// TIA Portal project "ESTHER_Gas_v4.0_4" (V13) (continued)
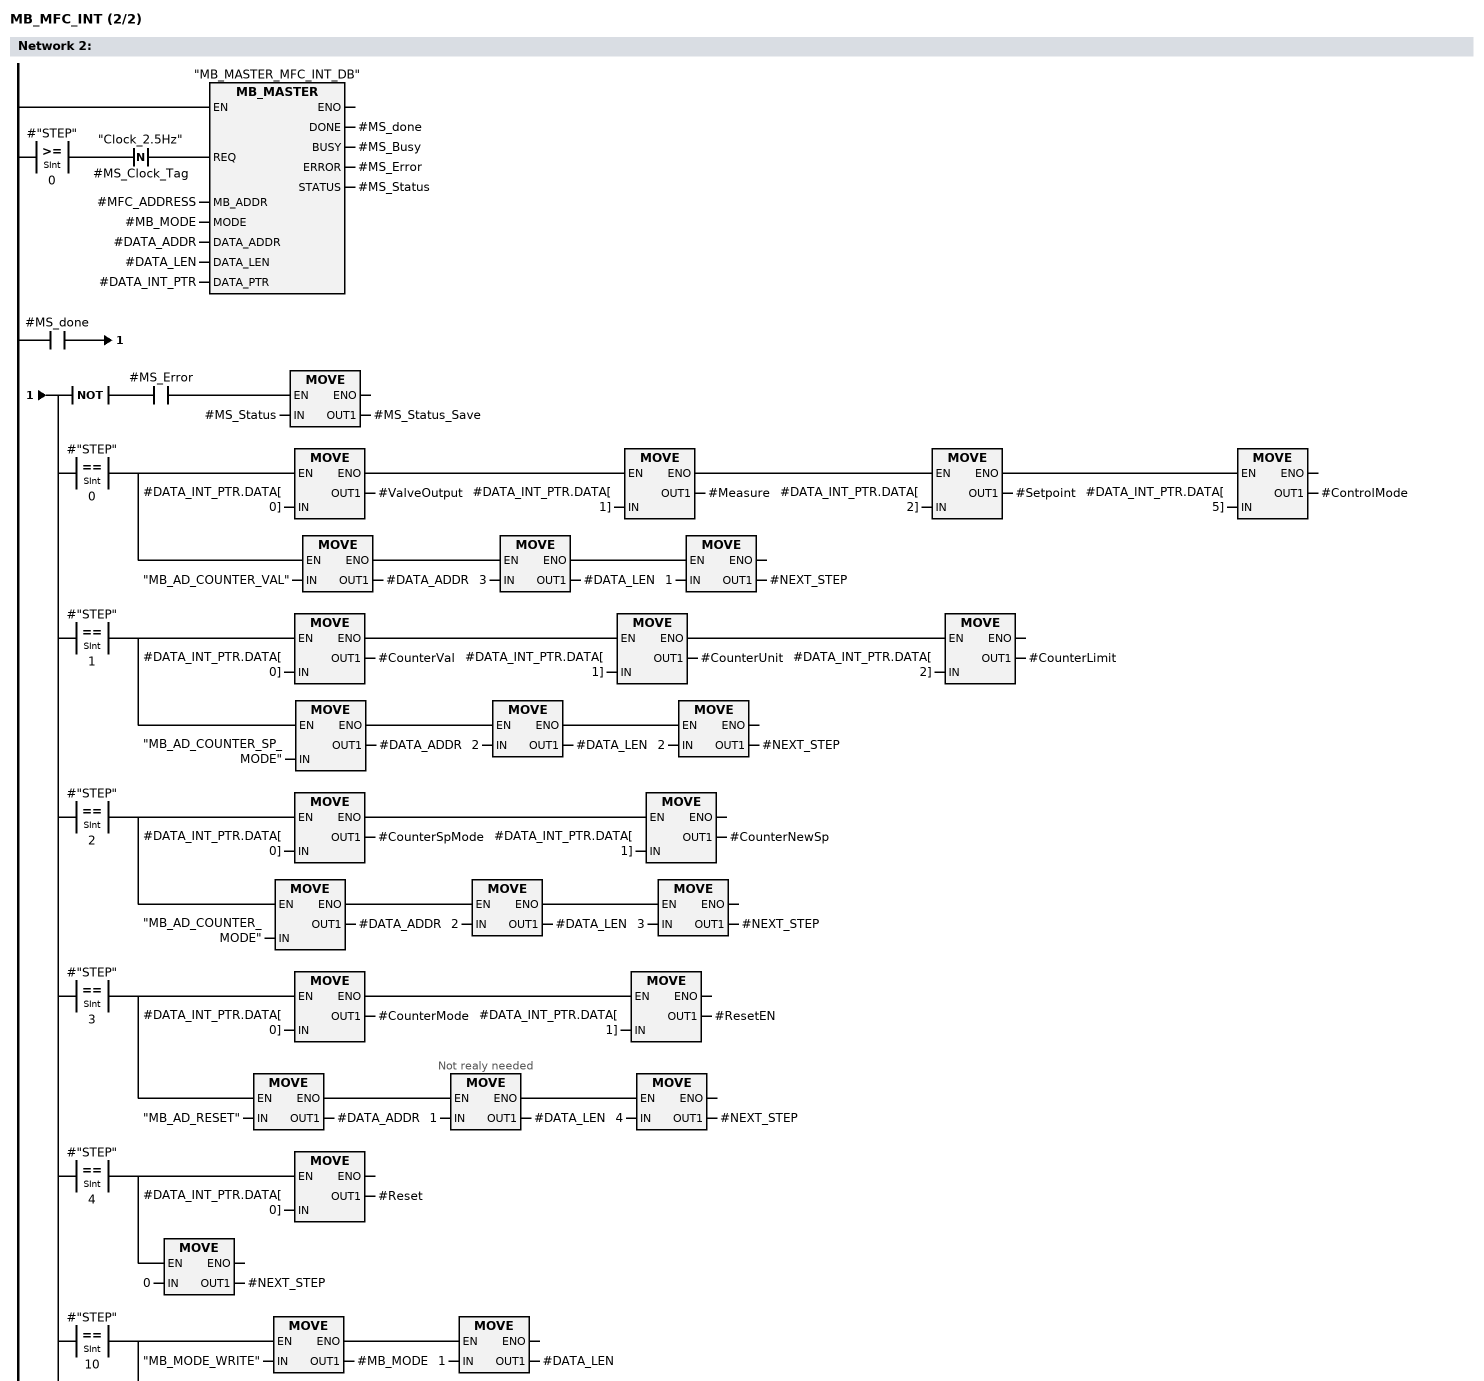
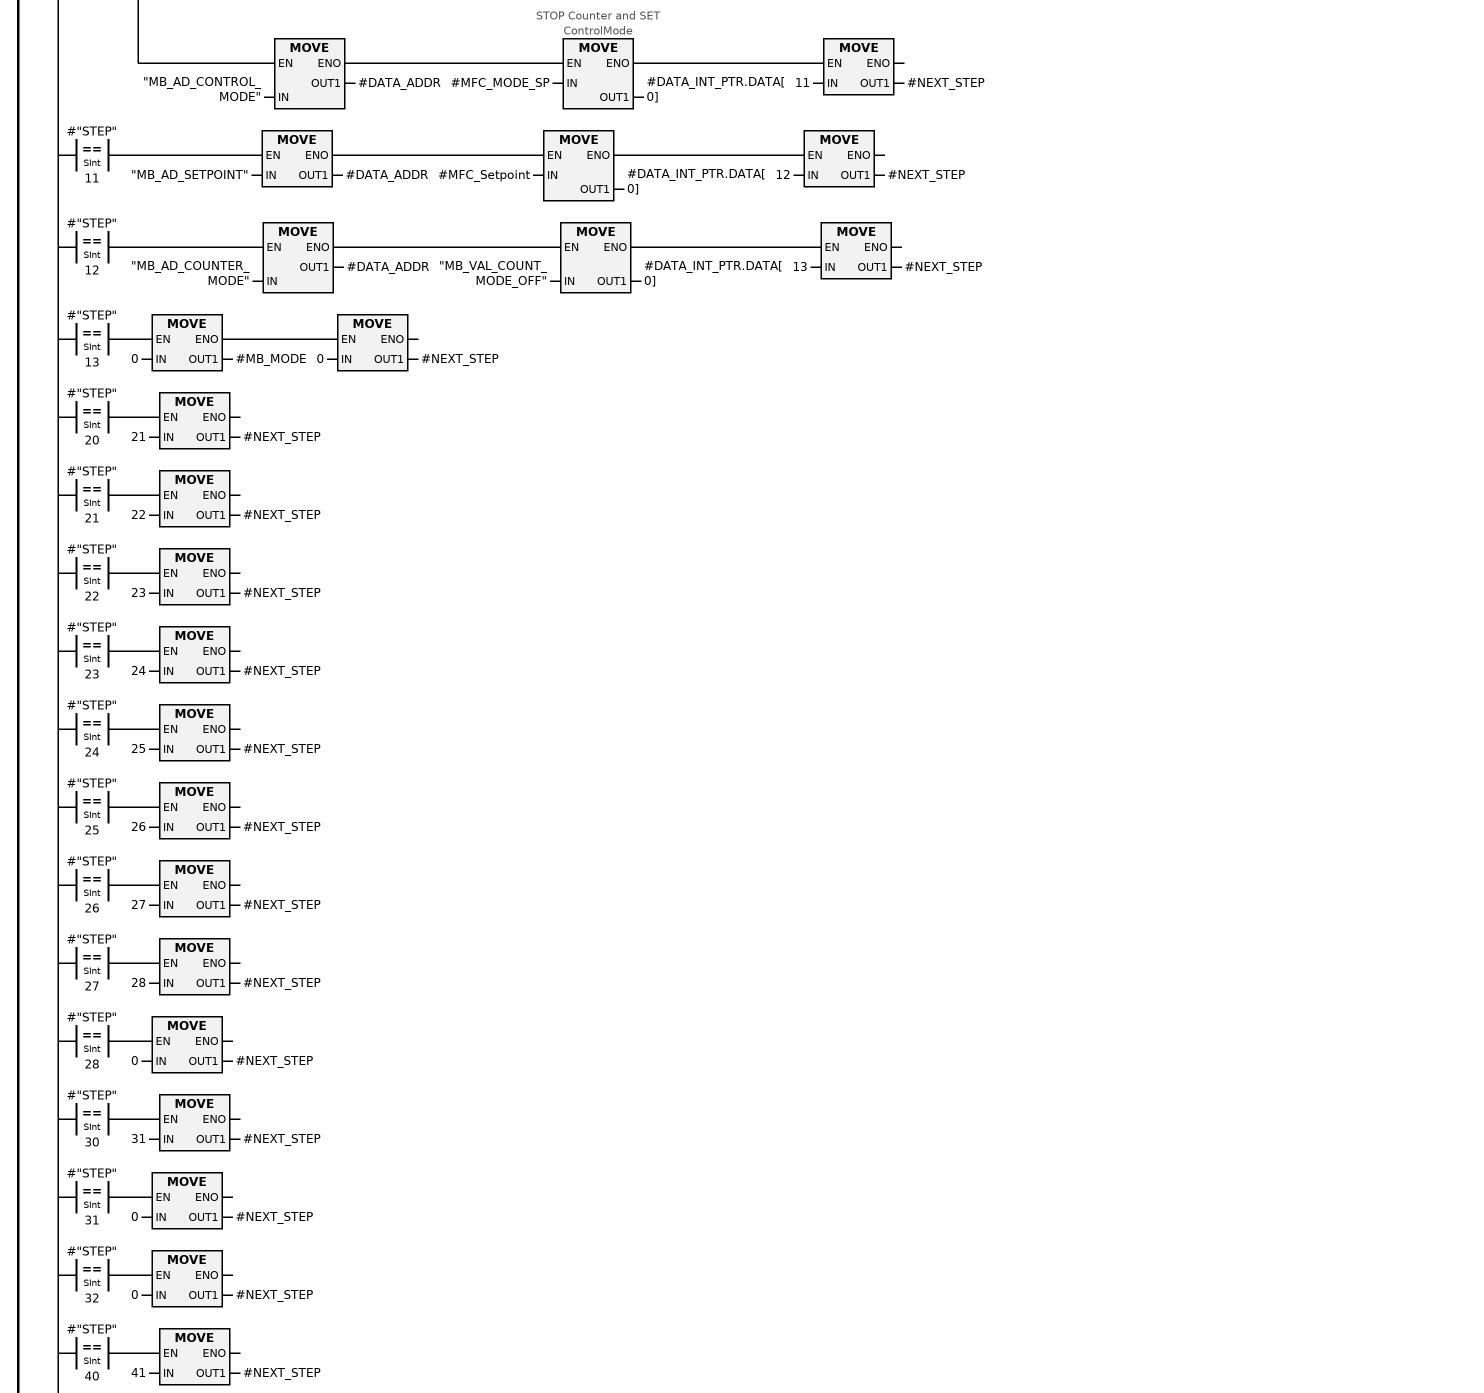
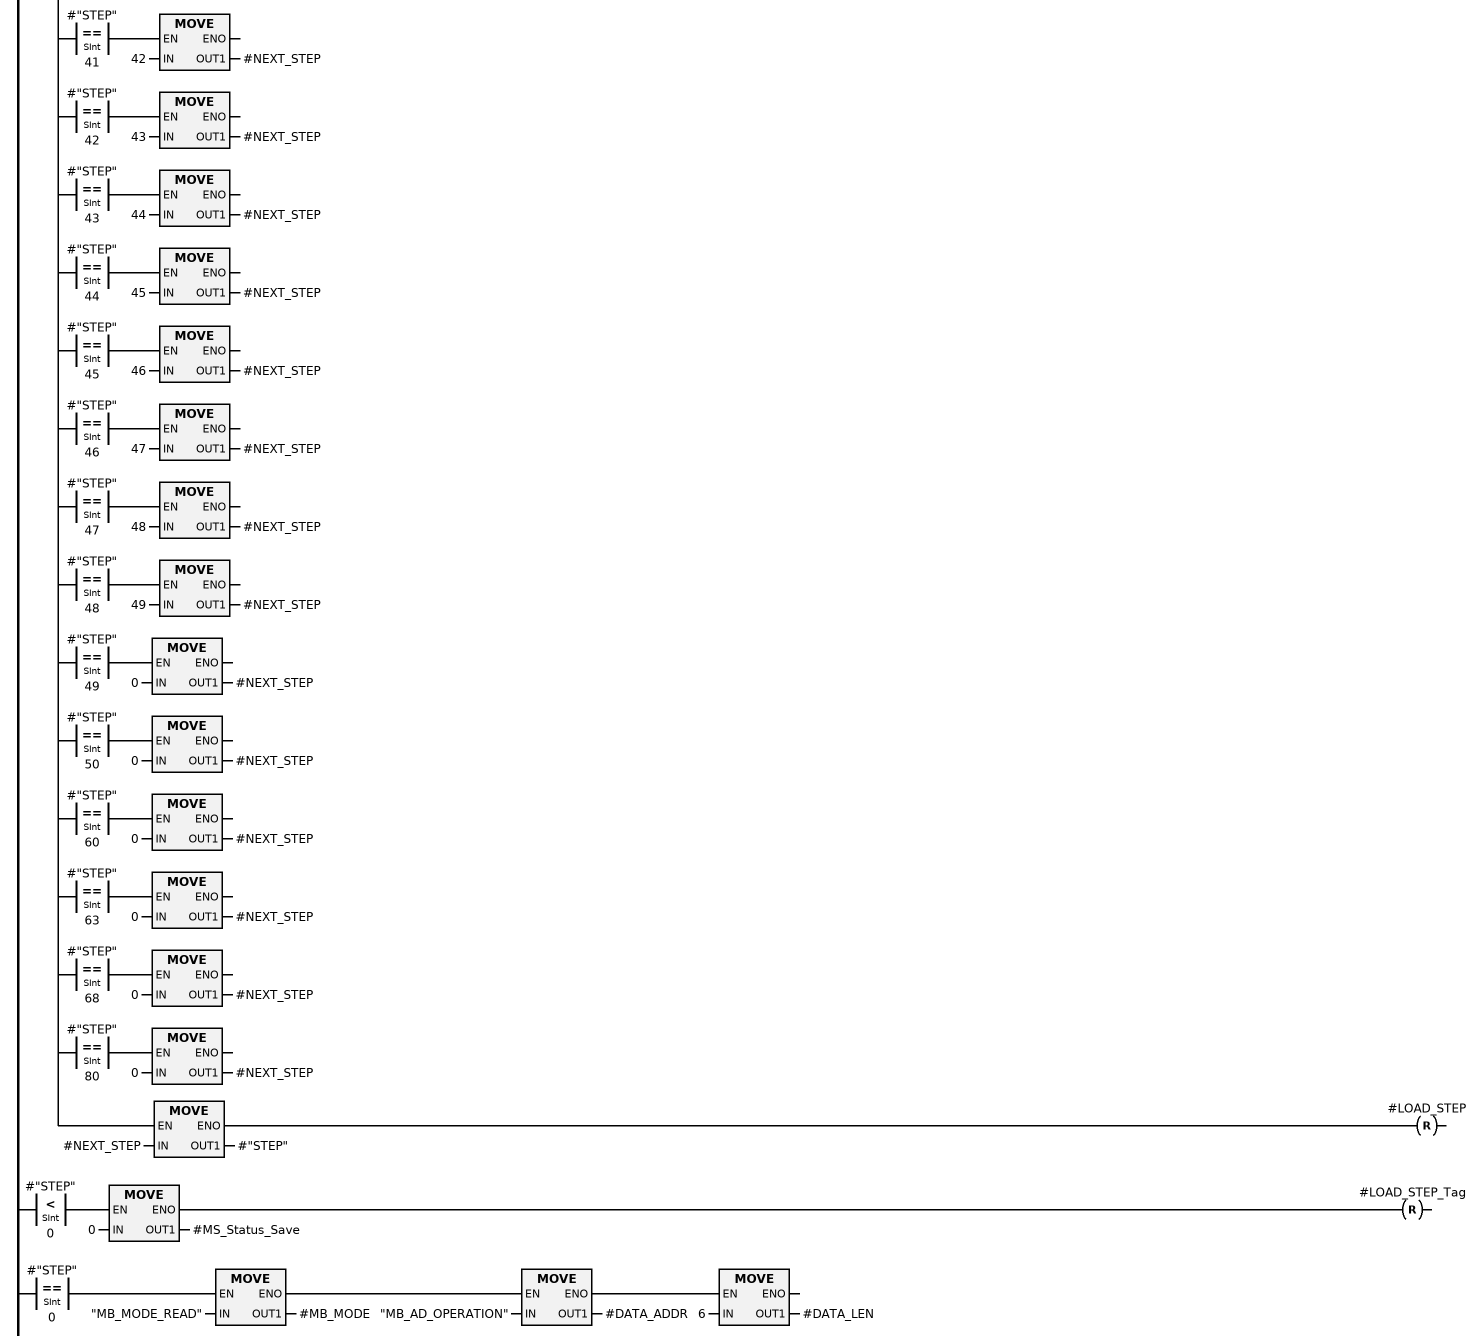
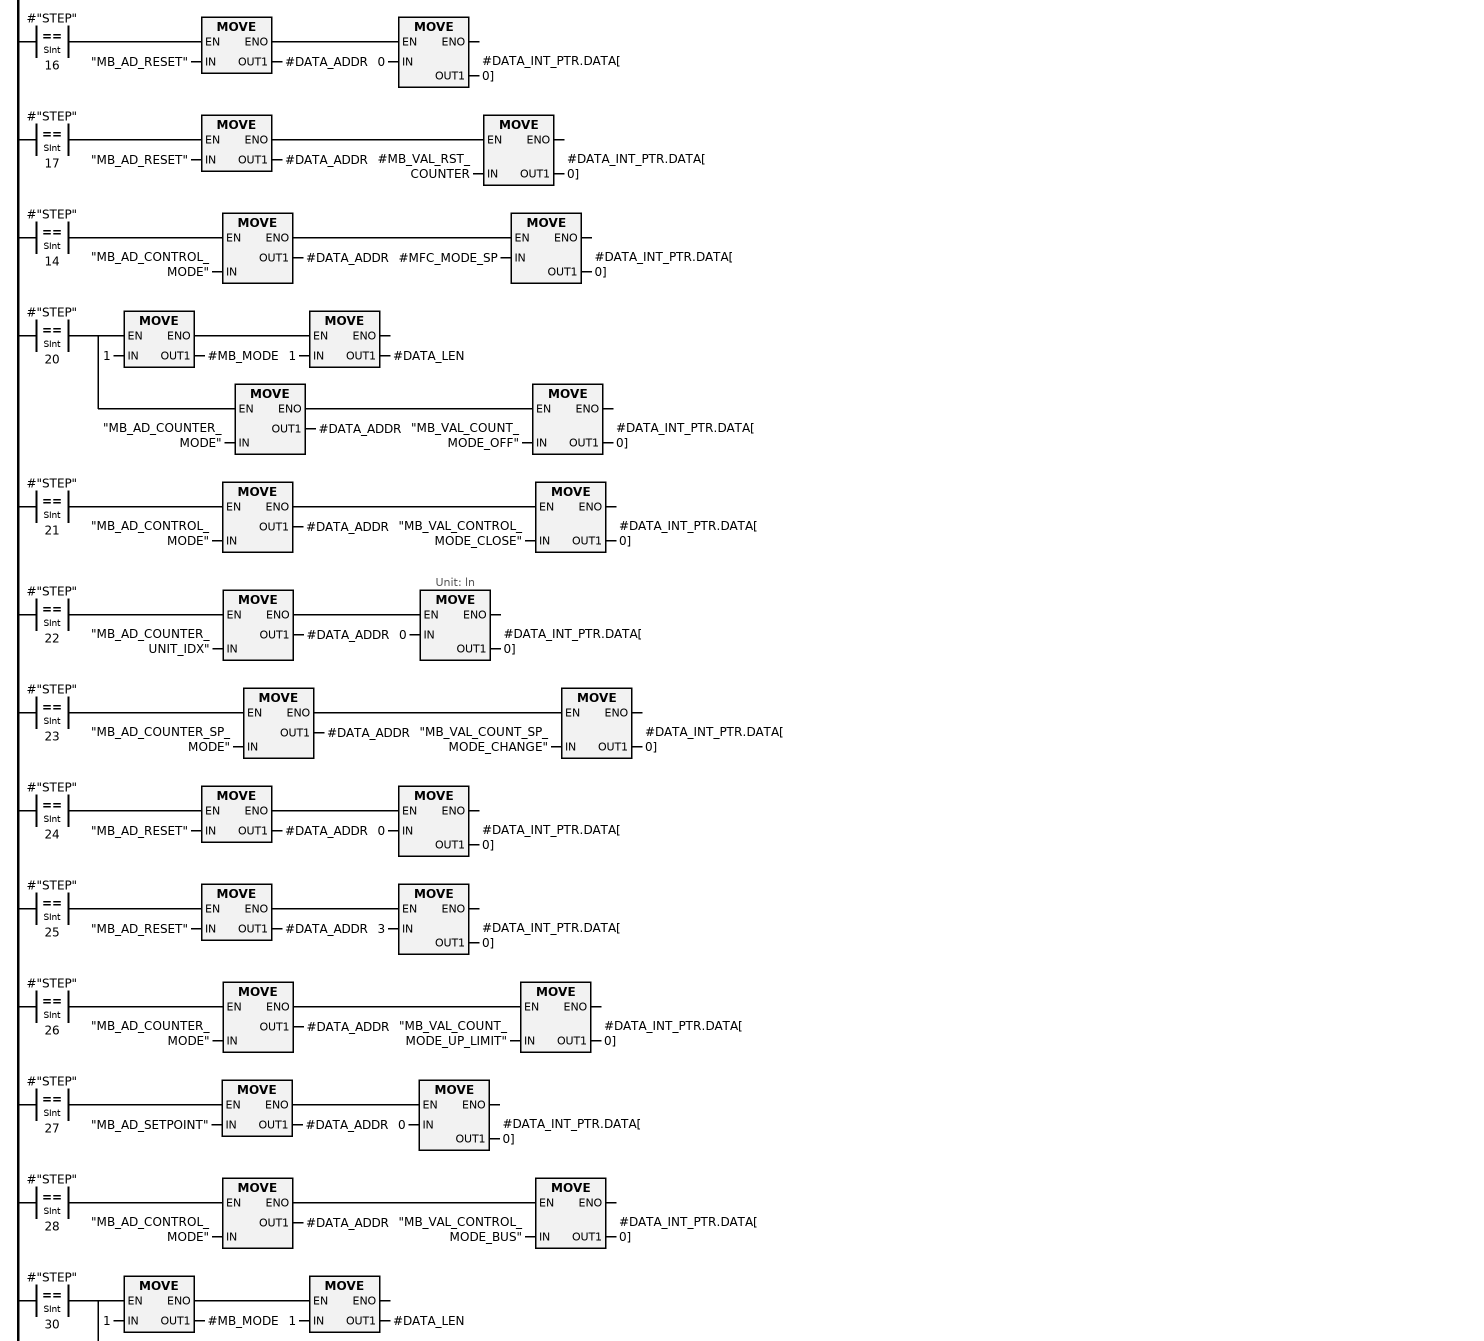
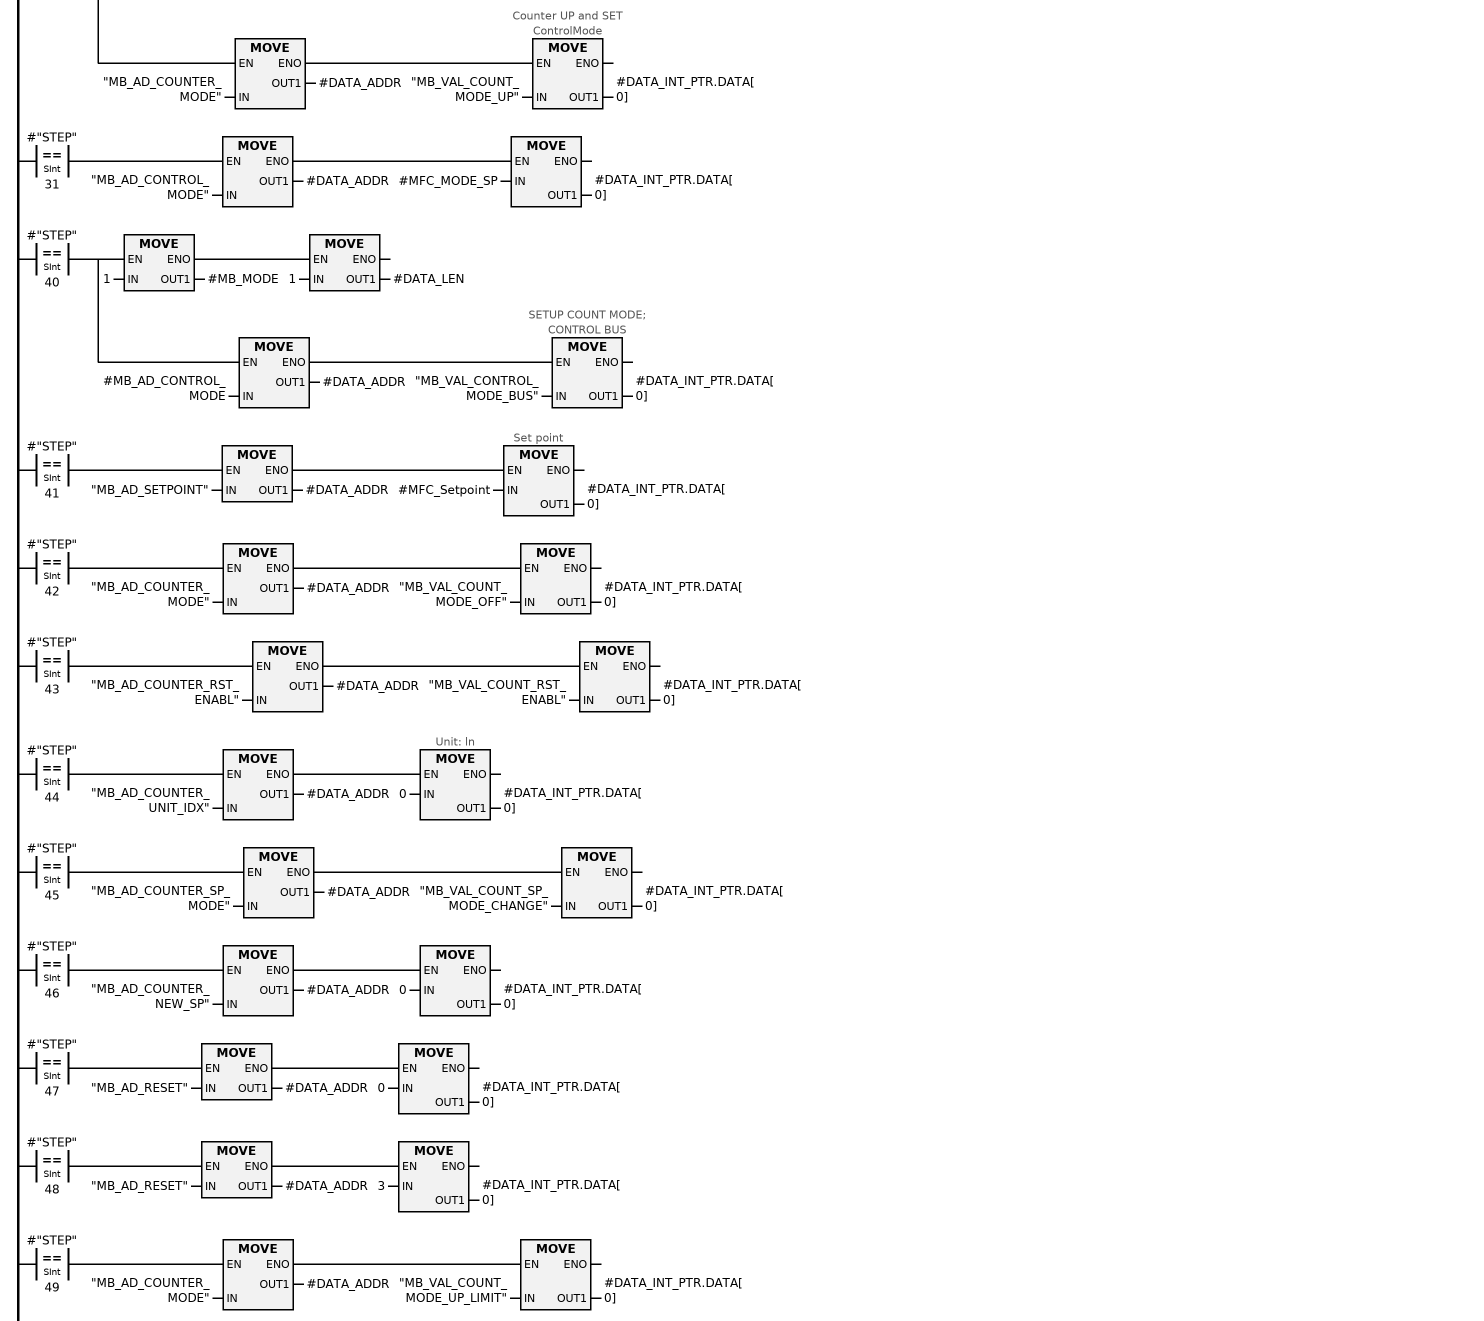
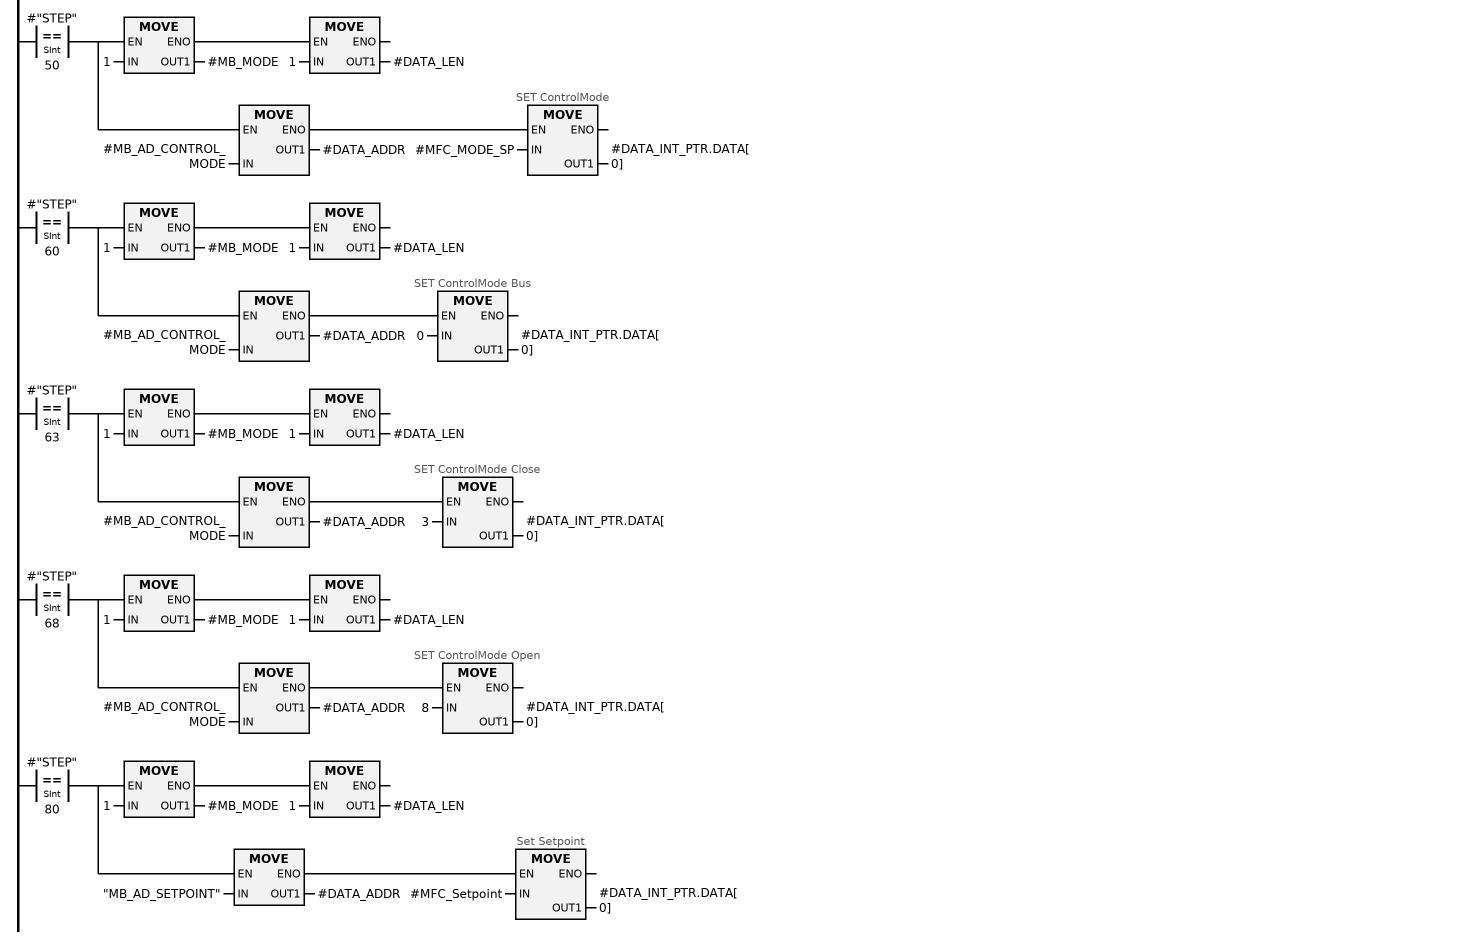
   #_w1 := (#"STEP" >= 0) AND NOT "Clock_2.5Hz" AND #MS_Clock_Tag;   // falling edge of "Clock_2.5Hz"
   #MS_Clock_Tag := "Clock_2.5Hz";
   "MB_MASTER_MFC_INT_DB"(REQ := #_w1,   // MB_MASTER
                          MB_ADDR := #MFC_ADDRESS,
                          MODE := #MB_MODE,
                          DATA_ADDR := #DATA_ADDR,
                          DATA_LEN := #DATA_LEN,
                          DATA_PTR := #DATA_INT_PTR,
                          DONE => #MS_done,
                          BUSY => #MS_Busy,
                          ERROR => #MS_Error,
                          STATUS => #MS_Status);
   IF NOT #MS_done AND #MS_Error THEN #MS_Status_Save := #MS_Status; END_IF;
   IF #MS_done AND (#"STEP" = 0) THEN
       #ValveOutput := #DATA_INT_PTR.DATA[0];
       #Measure := #DATA_INT_PTR.DATA[1];
       #Setpoint := #DATA_INT_PTR.DATA[2];
       #ControlMode := #DATA_INT_PTR.DATA[5];
       #DATA_ADDR := "MB_AD_COUNTER_VAL";
       #DATA_LEN := 3;
       #NEXT_STEP := 1;
   END_IF;
   IF #MS_done AND (#"STEP" = 1) THEN
       #CounterVal := #DATA_INT_PTR.DATA[0];
       #CounterUnit := #DATA_INT_PTR.DATA[1];
       #CounterLimit := #DATA_INT_PTR.DATA[2];
       #DATA_ADDR := "MB_AD_COUNTER_SP_MODE";
       #DATA_LEN := 2;
       #NEXT_STEP := 2;
   END_IF;
   IF #MS_done AND (#"STEP" = 2) THEN
       #CounterSpMode := #DATA_INT_PTR.DATA[0];
       #CounterNewSp := #DATA_INT_PTR.DATA[1];
       #DATA_ADDR := "MB_AD_COUNTER_MODE";
       #DATA_LEN := 2;
       #NEXT_STEP := 3;
   END_IF;
   IF #MS_done AND (#"STEP" = 3) THEN
       #CounterMode := #DATA_INT_PTR.DATA[0];
       #ResetEN := #DATA_INT_PTR.DATA[1];
       #DATA_ADDR := "MB_AD_RESET";
       #DATA_LEN := 1;   // Not realy needed
       #NEXT_STEP := 4;
   END_IF;
   IF #MS_done AND (#"STEP" = 4) THEN
       #Reset := #DATA_INT_PTR.DATA[0];
       #NEXT_STEP := 0;
   END_IF;
   IF #MS_done AND (#"STEP" = 10) THEN
       #MB_MODE := "MB_MODE_WRITE";
       #DATA_LEN := 1;
       #DATA_ADDR := "MB_AD_CONTROL_MODE";
       #DATA_INT_PTR.DATA[0] := #MFC_MODE_SP;   // STOP Counter and SET ControlMode
       #NEXT_STEP := 11;
   END_IF;
   IF #MS_done AND (#"STEP" = 11) THEN
       #DATA_ADDR := "MB_AD_SETPOINT";
       #DATA_INT_PTR.DATA[0] := #MFC_Setpoint;
       #NEXT_STEP := 12;
   END_IF;
   IF #MS_done AND (#"STEP" = 12) THEN
       #DATA_ADDR := "MB_AD_COUNTER_MODE";
       #DATA_INT_PTR.DATA[0] := "MB_VAL_COUNT_MODE_OFF";
       #NEXT_STEP := 13;
   END_IF;
   IF #MS_done AND (#"STEP" = 13) THEN
       #MB_MODE := 0;
       #NEXT_STEP := 0;
   END_IF;
   IF #MS_done AND (#"STEP" = 20) THEN #NEXT_STEP := 21; END_IF;
   IF #MS_done AND (#"STEP" = 21) THEN #NEXT_STEP := 22; END_IF;
   IF #MS_done AND (#"STEP" = 22) THEN #NEXT_STEP := 23; END_IF;
   IF #MS_done AND (#"STEP" = 23) THEN #NEXT_STEP := 24; END_IF;
   IF #MS_done AND (#"STEP" = 24) THEN #NEXT_STEP := 25; END_IF;
   IF #MS_done AND (#"STEP" = 25) THEN #NEXT_STEP := 26; END_IF;
   IF #MS_done AND (#"STEP" = 26) THEN #NEXT_STEP := 27; END_IF;
   IF #MS_done AND (#"STEP" = 27) THEN #NEXT_STEP := 28; END_IF;
   IF #MS_done AND (#"STEP" = 28) THEN #NEXT_STEP := 0; END_IF;
   IF #MS_done AND (#"STEP" = 30) THEN #NEXT_STEP := 31; END_IF;
   IF #MS_done AND (#"STEP" = 31) THEN #NEXT_STEP := 0; END_IF;
   IF #MS_done AND (#"STEP" = 32) THEN #NEXT_STEP := 0; END_IF;
   IF #MS_done AND (#"STEP" = 40) THEN #NEXT_STEP := 41; END_IF;
   IF #MS_done AND (#"STEP" = 41) THEN #NEXT_STEP := 42; END_IF;
   IF #MS_done AND (#"STEP" = 42) THEN #NEXT_STEP := 43; END_IF;
   IF #MS_done AND (#"STEP" = 43) THEN #NEXT_STEP := 44; END_IF;
   IF #MS_done AND (#"STEP" = 44) THEN #NEXT_STEP := 45; END_IF;
   IF #MS_done AND (#"STEP" = 45) THEN #NEXT_STEP := 46; END_IF;
   IF #MS_done AND (#"STEP" = 46) THEN #NEXT_STEP := 47; END_IF;
   IF #MS_done AND (#"STEP" = 47) THEN #NEXT_STEP := 48; END_IF;
   IF #MS_done AND (#"STEP" = 48) THEN #NEXT_STEP := 49; END_IF;
   IF #MS_done AND (#"STEP" = 49) THEN #NEXT_STEP := 0; END_IF;
   IF #MS_done AND (#"STEP" = 50) THEN #NEXT_STEP := 0; END_IF;
   IF #MS_done AND (#"STEP" = 60) THEN #NEXT_STEP := 0; END_IF;
   IF #MS_done AND (#"STEP" = 63) THEN #NEXT_STEP := 0; END_IF;
   IF #MS_done AND (#"STEP" = 68) THEN #NEXT_STEP := 0; END_IF;
   IF #MS_done AND (#"STEP" = 80) THEN #NEXT_STEP := 0; END_IF;
   IF #MS_done THEN
       #"STEP" := #NEXT_STEP;
       #LOAD_STEP := FALSE;
   END_IF;
   IF #"STEP" < 0 THEN
       #MS_Status_Save := 0;
       #LOAD_STEP_Tag := FALSE;
   END_IF;
   IF #"STEP" = 0 THEN
       #MB_MODE := "MB_MODE_READ";
       #DATA_ADDR := "MB_AD_OPERATION";
       #DATA_LEN := 6;
   END_IF;
   IF #"STEP" = 16 THEN
       #DATA_ADDR := "MB_AD_RESET";
       #DATA_INT_PTR.DATA[0] := 0;
   END_IF;
   IF #"STEP" = 17 THEN
       #DATA_ADDR := "MB_AD_RESET";
       #DATA_INT_PTR.DATA[0] := #MB_VAL_RST_COUNTER;
   END_IF;
   IF #"STEP" = 14 THEN
       #DATA_ADDR := "MB_AD_CONTROL_MODE";
       #DATA_INT_PTR.DATA[0] := #MFC_MODE_SP;
   END_IF;
   IF #"STEP" = 20 THEN
       #MB_MODE := 1;
       #DATA_LEN := 1;
       #DATA_ADDR := "MB_AD_COUNTER_MODE";
       #DATA_INT_PTR.DATA[0] := "MB_VAL_COUNT_MODE_OFF";
   END_IF;
   IF #"STEP" = 21 THEN
       #DATA_ADDR := "MB_AD_CONTROL_MODE";
       #DATA_INT_PTR.DATA[0] := "MB_VAL_CONTROL_MODE_CLOSE";
   END_IF;
   IF #"STEP" = 22 THEN
       #DATA_ADDR := "MB_AD_COUNTER_UNIT_IDX";
       #DATA_INT_PTR.DATA[0] := 0;   // Unit: ln
   END_IF;
   IF #"STEP" = 23 THEN
       #DATA_ADDR := "MB_AD_COUNTER_SP_MODE";
       #DATA_INT_PTR.DATA[0] := "MB_VAL_COUNT_SP_MODE_CHANGE";
   END_IF;
   IF #"STEP" = 24 THEN
       #DATA_ADDR := "MB_AD_RESET";
       #DATA_INT_PTR.DATA[0] := 0;
   END_IF;
   IF #"STEP" = 25 THEN
       #DATA_ADDR := "MB_AD_RESET";
       #DATA_INT_PTR.DATA[0] := 3;
   END_IF;
   IF #"STEP" = 26 THEN
       #DATA_ADDR := "MB_AD_COUNTER_MODE";
       #DATA_INT_PTR.DATA[0] := "MB_VAL_COUNT_MODE_UP_LIMIT";
   END_IF;
   IF #"STEP" = 27 THEN
       #DATA_ADDR := "MB_AD_SETPOINT";
       #DATA_INT_PTR.DATA[0] := 0;
   END_IF;
   IF #"STEP" = 28 THEN
       #DATA_ADDR := "MB_AD_CONTROL_MODE";
       #DATA_INT_PTR.DATA[0] := "MB_VAL_CONTROL_MODE_BUS";
   END_IF;
   IF #"STEP" = 30 THEN
       #MB_MODE := 1;
       #DATA_LEN := 1;
       #DATA_ADDR := "MB_AD_COUNTER_MODE";
       #DATA_INT_PTR.DATA[0] := "MB_VAL_COUNT_MODE_UP";   // Counter UP and SET ControlMode
   END_IF;
   IF #"STEP" = 31 THEN
       #DATA_ADDR := "MB_AD_CONTROL_MODE";
       #DATA_INT_PTR.DATA[0] := #MFC_MODE_SP;
   END_IF;
   IF #"STEP" = 40 THEN
       #MB_MODE := 1;
       #DATA_LEN := 1;
       #DATA_ADDR := #MB_AD_CONTROL_MODE;
       #DATA_INT_PTR.DATA[0] := "MB_VAL_CONTROL_MODE_BUS";   // SETUP COUNT MODE; CONTROL BUS
   END_IF;
   IF #"STEP" = 41 THEN
       #DATA_ADDR := "MB_AD_SETPOINT";
       #DATA_INT_PTR.DATA[0] := #MFC_Setpoint;   // Set point
   END_IF;
   IF #"STEP" = 42 THEN
       #DATA_ADDR := "MB_AD_COUNTER_MODE";
       #DATA_INT_PTR.DATA[0] := "MB_VAL_COUNT_MODE_OFF";
   END_IF;
   IF #"STEP" = 43 THEN